VERSION : 0.1
   VAR
      "1#炉体循环水泵电动阀" : "阀门_MODEL";
      "2#炉体循环水泵电动阀" : "阀门_MODEL";
      "3#炉体循环水泵电动阀" : "阀门_MODEL";
      "1#电极循环水泵电动阀" : "阀门_MODEL";
      "2#电极循环水泵电动阀" : "阀门_MODEL";
      "3#电极循环水泵电动阀" : "阀门_MODEL";
      "4#电极循环水泵电动阀" : "阀门_MODEL";
      "1#净环热水泵电动阀" : "阀门_MODEL";
      "2#净环热水泵电动阀" : "阀门_MODEL";
      "3#净环热水泵电动阀" : "阀门_MODEL";
      "4#净环热水泵电动阀" : "阀门_MODEL";
      "5#净环热水泵电动阀" : "阀门_MODEL";
      "1#浊环热水泵电动阀" : "阀门_MODEL";
      "2#浊环热水泵电动阀" : "阀门_MODEL";
      "3#浊环热水泵电动阀" : "阀门_MODEL";
      "4#浊环热水泵电动阀" : "阀门_MODEL";
      "5#浊环热水泵电动阀" : "阀门_MODEL";
      "6#浊环热水泵电动阀" : "阀门_MODEL";
      "7#浊环热水泵电动阀" : "阀门_MODEL";
      "8#浊环热水泵电动阀" : "阀门_MODEL";
      "1#冲渣泵电动阀" : "阀门_MODEL";
      "2#冲渣泵电动阀" : "阀门_MODEL";
      "3#冲渣泵电动阀" : "阀门_MODEL";
      "4#冲渣泵电动阀" : "阀门_MODEL";
      "5#冲渣泵电动阀" : "阀门_MODEL";
      "6#冲渣泵电动阀" : "阀门_MODEL";
      "7#冲渣泵电动阀" : "阀门_MODEL";
      "8#冲渣泵电动阀" : "阀门_MODEL";
      "1#柴油泵电动阀" : "阀门_MODEL";
      "2#柴油泵电动阀" : "阀门_MODEL";
      窑冷却泵电动阀 : "阀门_MODEL";
      Static4_1 : "阀门_MODEL";
      Static5_1 : "阀门_MODEL";
      Static6_1 : "阀门_MODEL";
      Static7_1 : "阀门_MODEL";
      Static8_1 : "阀门_MODEL";
      Static9_1 : "阀门_MODEL";
      Static10_1 : "阀门_MODEL";
      Static11_1 : "阀门_MODEL";
      Static12_1 : "阀门_MODEL";
      Static13_1 : "阀门_MODEL";
      Static14_1 : "阀门_MODEL";
      Static15_1 : "阀门_MODEL";
      Static16_1 : "阀门_MODEL";
      Static17_1 : "阀门_MODEL";
      Static18_1 : "阀门_MODEL";
      Static19_1 : "阀门_MODEL";
      Static20_1 : "阀门_MODEL";
      Static21_1 : "阀门_MODEL";
      Static22_1 : "阀门_MODEL";
      Static23_1 : "阀门_MODEL";
      Static24_1 : "阀门_MODEL";
      Static25_1 : "阀门_MODEL";
      Static26_1 : "阀门_MODEL";
      Static27_1 : "阀门_MODEL";
      Static28_1 : "阀门_MODEL";
      Static29_1 : "阀门_MODEL";
      Static30_1 : "阀门_MODEL";
      Static31_1 : "阀门_MODEL";
      Static32_1 : "阀门_MODEL";
      Static33_1 : "阀门_MODEL";
      Static34_1 : "阀门_MODEL";
      Static35_1 : "阀门_MODEL";
      Static36_1 : "阀门_MODEL";
      Static37_1 : "阀门_MODEL";
      Static38_1 : "阀门_MODEL";
      Static39_1 : "阀门_MODEL";
      Static40_1 : "阀门_MODEL";
      Static41_1 : "阀门_MODEL";
      Static42_1 : "阀门_MODEL";
      Static43_1 : "阀门_MODEL";
      Static44_1 : "阀门_MODEL";
      Static45_1 : "阀门_MODEL";
      Static46_1 : "阀门_MODEL";
      Static47_1 : "阀门_MODEL";
      Static48_1 : "阀门_MODEL";
      Static49_1 : "阀门_MODEL";
      Static50_1 : "阀门_MODEL";
      Static51_1 : "阀门_MODEL";
      Static52_1 : "阀门_MODEL";
      Static53_1 : "阀门_MODEL";
      Static54_1 : "阀门_MODEL";
      Static55_1 : "阀门_MODEL";
      Static56_1 : "阀门_MODEL";
      Static57_1 : "阀门_MODEL";
      Static58_1 : "阀门_MODEL";
      Static59_1 : "阀门_MODEL";
      Static60_1 : "阀门_MODEL";
      Static61_1 : "阀门_MODEL";
      Static62 : "阀门_MODEL";
      Static63 : "阀门_MODEL";
      Static64 : "阀门_MODEL";
      Static65 : "阀门_MODEL";
      Static66 : "阀门_MODEL";
      Static67 : "阀门_MODEL";
      Static68 : "阀门_MODEL";
      Static69 : "阀门_MODEL";
      Static70 : "阀门_MODEL";
      Static71 : "阀门_MODEL";
      Static72 : "阀门_MODEL";
      Static73 : "阀门_MODEL";
      Static74 : "阀门_MODEL";
      阀门_MODEL_Instance : "阀门_MODEL";
   END_VAR
   VAR CONSTANT
      Static3 : Bool;
      Static4 : Bool;
      Static5 : Bool;
      Static6 : Bool;
      Static7 : Bool;
      Static8 : Bool;
      Static9 : Bool;
      Static10 : Bool;
      Static11 : Bool;
      Static12 : Bool;
      Static13 : Bool;
      Static14 : Bool;
      Static15 : Bool;
      Static16 : Bool;
      Static17 : Bool;
      Static18 : Bool;
      Static19 : Bool;
      Static20 : Bool;
      Static21 : Bool;
      Static22 : Bool;
      Static23 : Bool;
      Static24 : Bool;
      Static25 : Bool;
      Static26 : Bool;
      Static27 : Bool;
      Static28 : Bool;
      Static29 : Bool;
      Static30 : Bool;
      Static31 : Bool;
      Static32 : Bool;
      Static33 : Bool;
      Static34 : Bool;
      Static35 : Bool;
      Static36 : Bool;
      Static37 : Bool;
      Static38 : Bool;
      Static39 : Bool;
      Static40 : Bool;
      Static41 : Bool;
      Static42 : Bool;
      Static43 : Bool;
      Static44 : Bool;
      Static45 : Bool;
      Static46 : Bool;
      Static47 : Bool;
      Static48 : Bool;
      Static49 : Bool;
      Static50 : Bool;
      Static51 : Bool;
      Static52 : Bool;
      Static53 : Bool;
      Static54 : Bool;
      Static55 : Bool;
      Static56 : Bool;
      Static57 : Bool;
      Static58 : Bool;
      Static59 : Bool;
      Static60 : Bool;
      Static61 : Bool;
   END_VAR
BEGIN

REGION Network 1
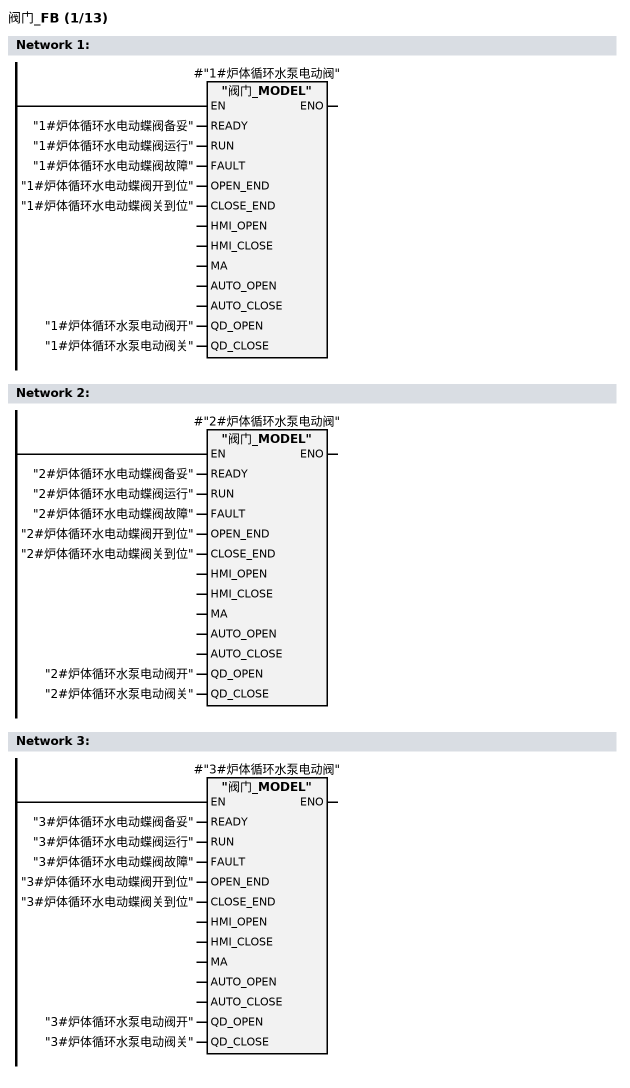
   RUNG wire#powerrail
      #"1#炉体循环水泵电动阀"(READY := "1#炉体循环水电动蝶阀备妥", RUN := "1#炉体循环水电动蝶阀运行", FAULT := "1#炉体循环水电动蝶阀故障", OPEN_END := "1#炉体循环水电动蝶阀开到位", CLOSE_END := "1#炉体循环水电动蝶阀关到位", HMI_OPEN :=, HMI_CLOSE :=, MA :=, AUTO_OPEN :=, AUTO_CLOSE :=, QD_OPEN := "1#炉体循环水泵电动阀开", QD_CLOSE := "1#炉体循环水泵电动阀关")
   END_RUNG
   // the same network as SCL:
   #"1#炉体循环水泵电动阀"(READY := "1#炉体循环水电动蝶阀备妥",   // "阀门_MODEL"
                  RUN := "1#炉体循环水电动蝶阀运行",
                  FAULT := "1#炉体循环水电动蝶阀故障",
                  OPEN_END := "1#炉体循环水电动蝶阀开到位",
                  CLOSE_END := "1#炉体循环水电动蝶阀关到位",
                  QD_OPEN := "1#炉体循环水泵电动阀开",
                  QD_CLOSE := "1#炉体循环水泵电动阀关");
END_REGION

REGION Network 2
   RUNG wire#powerrail
      #"2#炉体循环水泵电动阀"(READY := "2#炉体循环水电动蝶阀备妥", RUN := "2#炉体循环水电动蝶阀运行", FAULT := "2#炉体循环水电动蝶阀故障", OPEN_END := "2#炉体循环水电动蝶阀开到位", CLOSE_END := "2#炉体循环水电动蝶阀关到位", HMI_OPEN :=, HMI_CLOSE :=, MA :=, AUTO_OPEN :=, AUTO_CLOSE :=, QD_OPEN := "2#炉体循环水泵电动阀开", QD_CLOSE := "2#炉体循环水泵电动阀关")
   END_RUNG
   // the same network as SCL:
   #"2#炉体循环水泵电动阀"(READY := "2#炉体循环水电动蝶阀备妥",   // "阀门_MODEL"
                  RUN := "2#炉体循环水电动蝶阀运行",
                  FAULT := "2#炉体循环水电动蝶阀故障",
                  OPEN_END := "2#炉体循环水电动蝶阀开到位",
                  CLOSE_END := "2#炉体循环水电动蝶阀关到位",
                  QD_OPEN := "2#炉体循环水泵电动阀开",
                  QD_CLOSE := "2#炉体循环水泵电动阀关");
END_REGION

REGION Network 3
   RUNG wire#powerrail
      #"3#炉体循环水泵电动阀"(READY := "3#炉体循环水电动蝶阀备妥", RUN := "3#炉体循环水电动蝶阀运行", FAULT := "3#炉体循环水电动蝶阀故障", OPEN_END := "3#炉体循环水电动蝶阀开到位", CLOSE_END := "3#炉体循环水电动蝶阀关到位", HMI_OPEN :=, HMI_CLOSE :=, MA :=, AUTO_OPEN :=, AUTO_CLOSE :=, QD_OPEN := "3#炉体循环水泵电动阀开", QD_CLOSE := "3#炉体循环水泵电动阀关")
   END_RUNG
   // the same network as SCL:
   #"3#炉体循环水泵电动阀"(READY := "3#炉体循环水电动蝶阀备妥",   // "阀门_MODEL"
                  RUN := "3#炉体循环水电动蝶阀运行",
                  FAULT := "3#炉体循环水电动蝶阀故障",
                  OPEN_END := "3#炉体循环水电动蝶阀开到位",
                  CLOSE_END := "3#炉体循环水电动蝶阀关到位",
                  QD_OPEN := "3#炉体循环水泵电动阀开",
                  QD_CLOSE := "3#炉体循环水泵电动阀关");
END_REGION

REGION Network 4
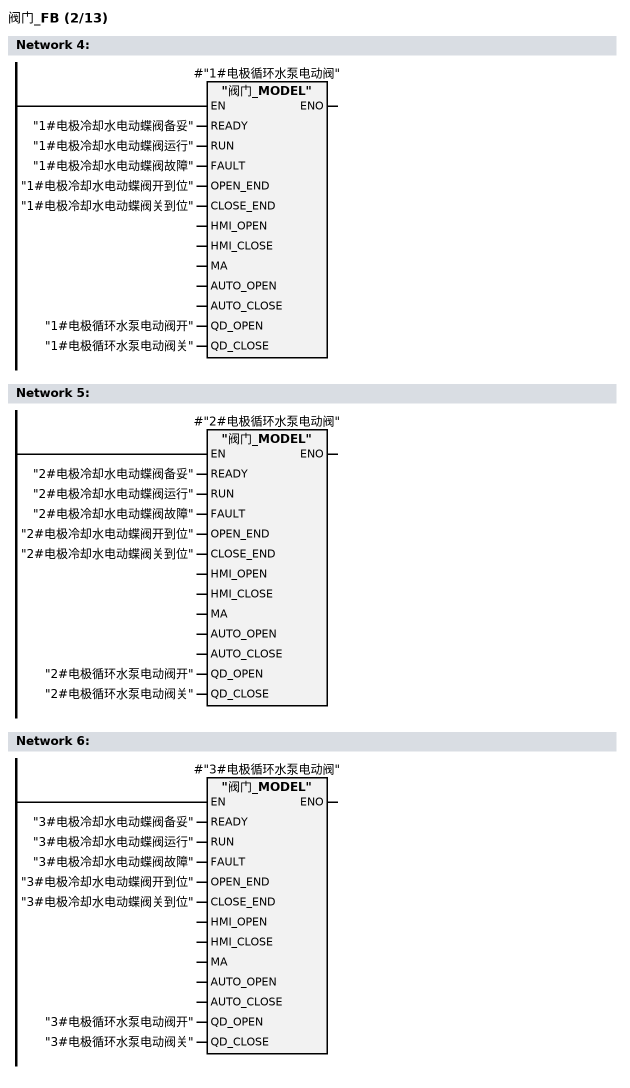
   RUNG wire#powerrail
      #"1#电极循环水泵电动阀"(READY := "1#电极冷却水电动蝶阀备妥", RUN := "1#电极冷却水电动蝶阀运行", FAULT := "1#电极冷却水电动蝶阀故障", OPEN_END := "1#电极冷却水电动蝶阀开到位", CLOSE_END := "1#电极冷却水电动蝶阀关到位", HMI_OPEN :=, HMI_CLOSE :=, MA :=, AUTO_OPEN :=, AUTO_CLOSE :=, QD_OPEN := "1#电极循环水泵电动阀开", QD_CLOSE := "1#电极循环水泵电动阀关")
   END_RUNG
   // the same network as SCL:
   #"1#电极循环水泵电动阀"(READY := "1#电极冷却水电动蝶阀备妥",   // "阀门_MODEL"
                  RUN := "1#电极冷却水电动蝶阀运行",
                  FAULT := "1#电极冷却水电动蝶阀故障",
                  OPEN_END := "1#电极冷却水电动蝶阀开到位",
                  CLOSE_END := "1#电极冷却水电动蝶阀关到位",
                  QD_OPEN := "1#电极循环水泵电动阀开",
                  QD_CLOSE := "1#电极循环水泵电动阀关");
END_REGION

REGION Network 5
   RUNG wire#powerrail
      #"2#电极循环水泵电动阀"(READY := "2#电极冷却水电动蝶阀备妥", RUN := "2#电极冷却水电动蝶阀运行", FAULT := "2#电极冷却水电动蝶阀故障", OPEN_END := "2#电极冷却水电动蝶阀开到位", CLOSE_END := "2#电极冷却水电动蝶阀关到位", HMI_OPEN :=, HMI_CLOSE :=, MA :=, AUTO_OPEN :=, AUTO_CLOSE :=, QD_OPEN := "2#电极循环水泵电动阀开", QD_CLOSE := "2#电极循环水泵电动阀关")
   END_RUNG
   // the same network as SCL:
   #"2#电极循环水泵电动阀"(READY := "2#电极冷却水电动蝶阀备妥",   // "阀门_MODEL"
                  RUN := "2#电极冷却水电动蝶阀运行",
                  FAULT := "2#电极冷却水电动蝶阀故障",
                  OPEN_END := "2#电极冷却水电动蝶阀开到位",
                  CLOSE_END := "2#电极冷却水电动蝶阀关到位",
                  QD_OPEN := "2#电极循环水泵电动阀开",
                  QD_CLOSE := "2#电极循环水泵电动阀关");
END_REGION

REGION Network 6
   RUNG wire#powerrail
      #"3#电极循环水泵电动阀"(READY := "3#电极冷却水电动蝶阀备妥", RUN := "3#电极冷却水电动蝶阀运行", FAULT := "3#电极冷却水电动蝶阀故障", OPEN_END := "3#电极冷却水电动蝶阀开到位", CLOSE_END := "3#电极冷却水电动蝶阀关到位", HMI_OPEN :=, HMI_CLOSE :=, MA :=, AUTO_OPEN :=, AUTO_CLOSE :=, QD_OPEN := "3#电极循环水泵电动阀开", QD_CLOSE := "3#电极循环水泵电动阀关")
   END_RUNG
   // the same network as SCL:
   #"3#电极循环水泵电动阀"(READY := "3#电极冷却水电动蝶阀备妥",   // "阀门_MODEL"
                  RUN := "3#电极冷却水电动蝶阀运行",
                  FAULT := "3#电极冷却水电动蝶阀故障",
                  OPEN_END := "3#电极冷却水电动蝶阀开到位",
                  CLOSE_END := "3#电极冷却水电动蝶阀关到位",
                  QD_OPEN := "3#电极循环水泵电动阀开",
                  QD_CLOSE := "3#电极循环水泵电动阀关");
END_REGION

REGION Network 7
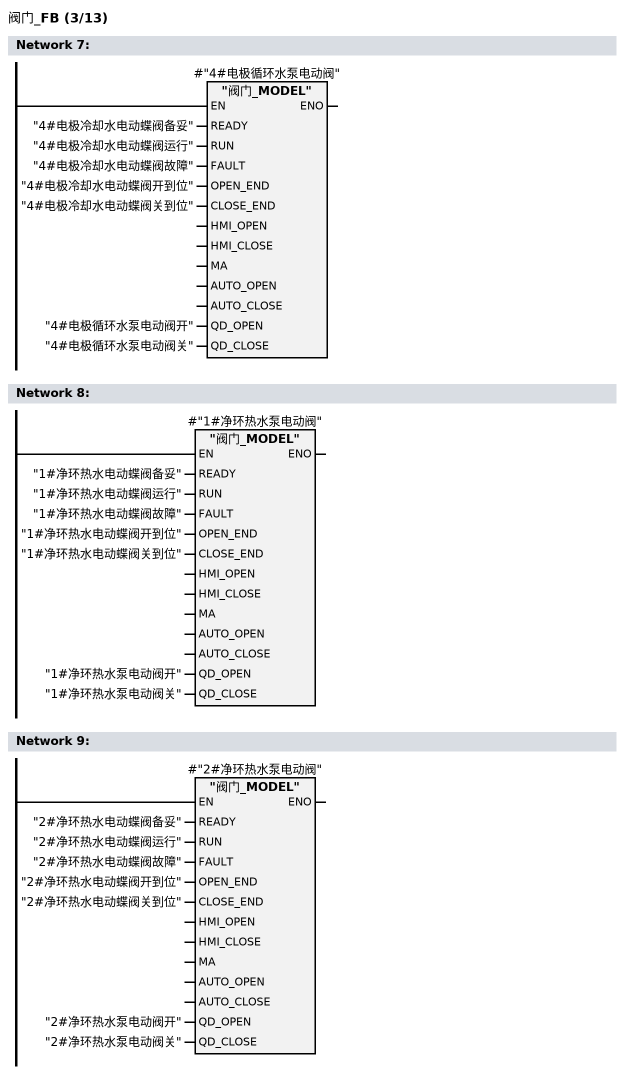
   RUNG wire#powerrail
      #"4#电极循环水泵电动阀"(READY := "4#电极冷却水电动蝶阀备妥", RUN := "4#电极冷却水电动蝶阀运行", FAULT := "4#电极冷却水电动蝶阀故障", OPEN_END := "4#电极冷却水电动蝶阀开到位", CLOSE_END := "4#电极冷却水电动蝶阀关到位", HMI_OPEN :=, HMI_CLOSE :=, MA :=, AUTO_OPEN :=, AUTO_CLOSE :=, QD_OPEN := "4#电极循环水泵电动阀开", QD_CLOSE := "4#电极循环水泵电动阀关")
   END_RUNG
   // the same network as SCL:
   #"4#电极循环水泵电动阀"(READY := "4#电极冷却水电动蝶阀备妥",   // "阀门_MODEL"
                  RUN := "4#电极冷却水电动蝶阀运行",
                  FAULT := "4#电极冷却水电动蝶阀故障",
                  OPEN_END := "4#电极冷却水电动蝶阀开到位",
                  CLOSE_END := "4#电极冷却水电动蝶阀关到位",
                  QD_OPEN := "4#电极循环水泵电动阀开",
                  QD_CLOSE := "4#电极循环水泵电动阀关");
END_REGION

REGION Network 8
   RUNG wire#powerrail
      #"1#净环热水泵电动阀"(READY := "1#净环热水电动蝶阀备妥", RUN := "1#净环热水电动蝶阀运行", FAULT := "1#净环热水电动蝶阀故障", OPEN_END := "1#净环热水电动蝶阀开到位", CLOSE_END := "1#净环热水电动蝶阀关到位", HMI_OPEN :=, HMI_CLOSE :=, MA :=, AUTO_OPEN :=, AUTO_CLOSE :=, QD_OPEN := "1#净环热水泵电动阀开", QD_CLOSE := "1#净环热水泵电动阀关")
   END_RUNG
   // the same network as SCL:
   #"1#净环热水泵电动阀"(READY := "1#净环热水电动蝶阀备妥",   // "阀门_MODEL"
                 RUN := "1#净环热水电动蝶阀运行",
                 FAULT := "1#净环热水电动蝶阀故障",
                 OPEN_END := "1#净环热水电动蝶阀开到位",
                 CLOSE_END := "1#净环热水电动蝶阀关到位",
                 QD_OPEN := "1#净环热水泵电动阀开",
                 QD_CLOSE := "1#净环热水泵电动阀关");
END_REGION

REGION Network 9
   RUNG wire#powerrail
      #"2#净环热水泵电动阀"(READY := "2#净环热水电动蝶阀备妥", RUN := "2#净环热水电动蝶阀运行", FAULT := "2#净环热水电动蝶阀故障", OPEN_END := "2#净环热水电动蝶阀开到位", CLOSE_END := "2#净环热水电动蝶阀关到位", HMI_OPEN :=, HMI_CLOSE :=, MA :=, AUTO_OPEN :=, AUTO_CLOSE :=, QD_OPEN := "2#净环热水泵电动阀开", QD_CLOSE := "2#净环热水泵电动阀关")
   END_RUNG
   // the same network as SCL:
   #"2#净环热水泵电动阀"(READY := "2#净环热水电动蝶阀备妥",   // "阀门_MODEL"
                 RUN := "2#净环热水电动蝶阀运行",
                 FAULT := "2#净环热水电动蝶阀故障",
                 OPEN_END := "2#净环热水电动蝶阀开到位",
                 CLOSE_END := "2#净环热水电动蝶阀关到位",
                 QD_OPEN := "2#净环热水泵电动阀开",
                 QD_CLOSE := "2#净环热水泵电动阀关");
END_REGION

REGION Network 10
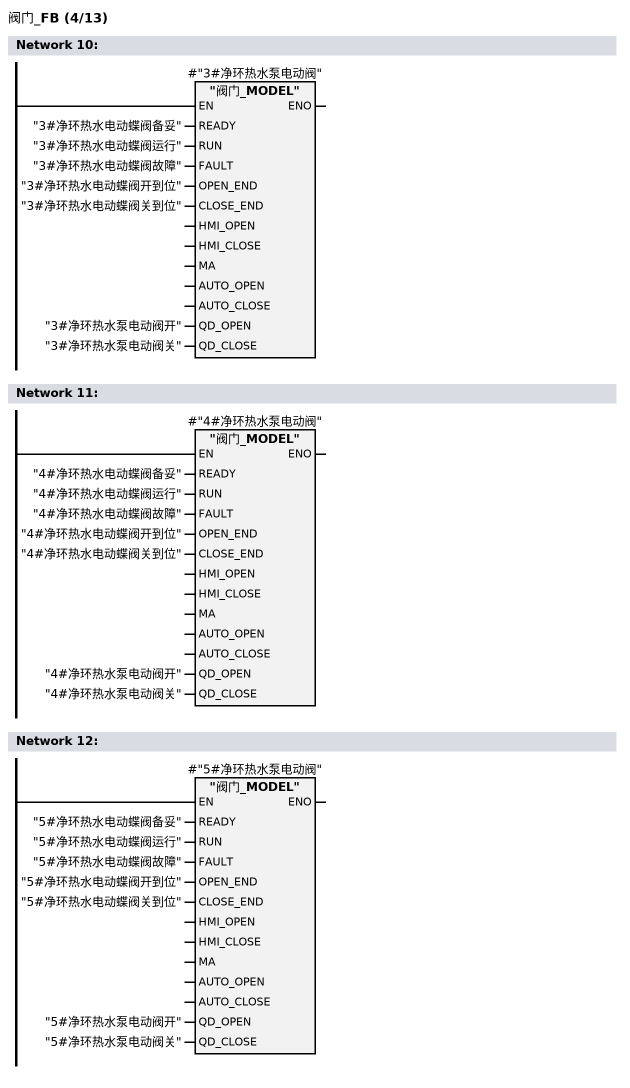
   RUNG wire#powerrail
      #"3#净环热水泵电动阀"(READY := "3#净环热水电动蝶阀备妥", RUN := "3#净环热水电动蝶阀运行", FAULT := "3#净环热水电动蝶阀故障", OPEN_END := "3#净环热水电动蝶阀开到位", CLOSE_END := "3#净环热水电动蝶阀关到位", HMI_OPEN :=, HMI_CLOSE :=, MA :=, AUTO_OPEN :=, AUTO_CLOSE :=, QD_OPEN := "3#净环热水泵电动阀开", QD_CLOSE := "3#净环热水泵电动阀关")
   END_RUNG
   // the same network as SCL:
   #"3#净环热水泵电动阀"(READY := "3#净环热水电动蝶阀备妥",   // "阀门_MODEL"
                 RUN := "3#净环热水电动蝶阀运行",
                 FAULT := "3#净环热水电动蝶阀故障",
                 OPEN_END := "3#净环热水电动蝶阀开到位",
                 CLOSE_END := "3#净环热水电动蝶阀关到位",
                 QD_OPEN := "3#净环热水泵电动阀开",
                 QD_CLOSE := "3#净环热水泵电动阀关");
END_REGION

REGION Network 11
   RUNG wire#powerrail
      #"4#净环热水泵电动阀"(READY := "4#净环热水电动蝶阀备妥", RUN := "4#净环热水电动蝶阀运行", FAULT := "4#净环热水电动蝶阀故障", OPEN_END := "4#净环热水电动蝶阀开到位", CLOSE_END := "4#净环热水电动蝶阀关到位", HMI_OPEN :=, HMI_CLOSE :=, MA :=, AUTO_OPEN :=, AUTO_CLOSE :=, QD_OPEN := "4#净环热水泵电动阀开", QD_CLOSE := "4#净环热水泵电动阀关")
   END_RUNG
   // the same network as SCL:
   #"4#净环热水泵电动阀"(READY := "4#净环热水电动蝶阀备妥",   // "阀门_MODEL"
                 RUN := "4#净环热水电动蝶阀运行",
                 FAULT := "4#净环热水电动蝶阀故障",
                 OPEN_END := "4#净环热水电动蝶阀开到位",
                 CLOSE_END := "4#净环热水电动蝶阀关到位",
                 QD_OPEN := "4#净环热水泵电动阀开",
                 QD_CLOSE := "4#净环热水泵电动阀关");
END_REGION

REGION Network 12
   RUNG wire#powerrail
      #"5#净环热水泵电动阀"(READY := "5#净环热水电动蝶阀备妥", RUN := "5#净环热水电动蝶阀运行", FAULT := "5#净环热水电动蝶阀故障", OPEN_END := "5#净环热水电动蝶阀开到位", CLOSE_END := "5#净环热水电动蝶阀关到位", HMI_OPEN :=, HMI_CLOSE :=, MA :=, AUTO_OPEN :=, AUTO_CLOSE :=, QD_OPEN := "5#净环热水泵电动阀开", QD_CLOSE := "5#净环热水泵电动阀关")
   END_RUNG
   // the same network as SCL:
   #"5#净环热水泵电动阀"(READY := "5#净环热水电动蝶阀备妥",   // "阀门_MODEL"
                 RUN := "5#净环热水电动蝶阀运行",
                 FAULT := "5#净环热水电动蝶阀故障",
                 OPEN_END := "5#净环热水电动蝶阀开到位",
                 CLOSE_END := "5#净环热水电动蝶阀关到位",
                 QD_OPEN := "5#净环热水泵电动阀开",
                 QD_CLOSE := "5#净环热水泵电动阀关");
END_REGION

REGION Network 13
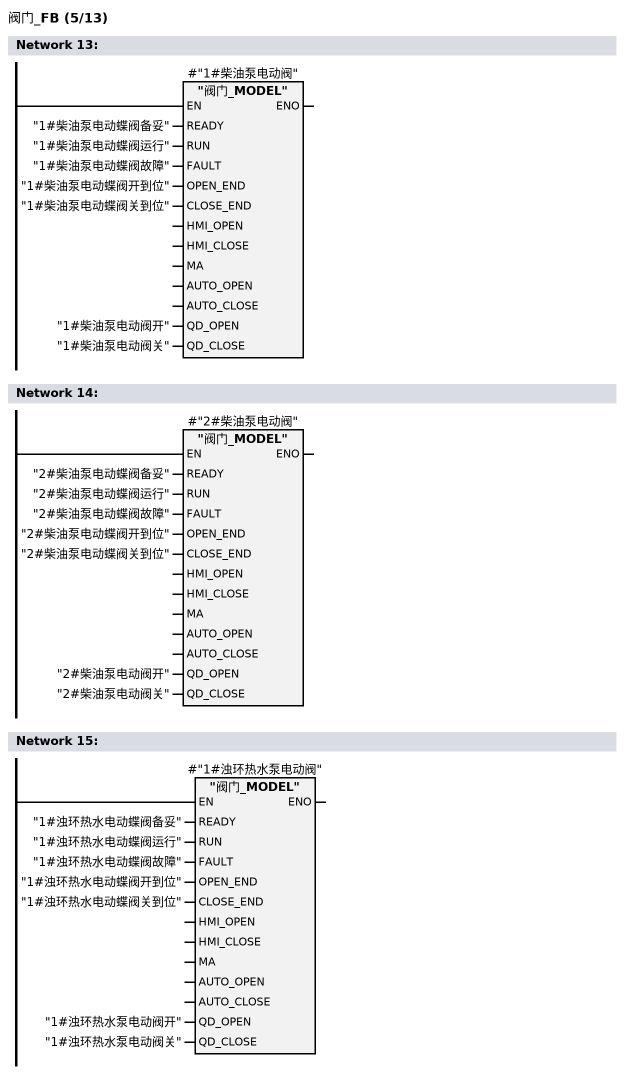
   RUNG wire#powerrail
      #"1#柴油泵电动阀"(READY := "1#柴油泵电动蝶阀备妥", RUN := "1#柴油泵电动蝶阀运行", FAULT := "1#柴油泵电动蝶阀故障", OPEN_END := "1#柴油泵电动蝶阀开到位", CLOSE_END := "1#柴油泵电动蝶阀关到位", HMI_OPEN :=, HMI_CLOSE :=, MA :=, AUTO_OPEN :=, AUTO_CLOSE :=, QD_OPEN := "1#柴油泵电动阀开", QD_CLOSE := "1#柴油泵电动阀关")
   END_RUNG
   // the same network as SCL:
   #"1#柴油泵电动阀"(READY := "1#柴油泵电动蝶阀备妥",   // "阀门_MODEL"
               RUN := "1#柴油泵电动蝶阀运行",
               FAULT := "1#柴油泵电动蝶阀故障",
               OPEN_END := "1#柴油泵电动蝶阀开到位",
               CLOSE_END := "1#柴油泵电动蝶阀关到位",
               QD_OPEN := "1#柴油泵电动阀开",
               QD_CLOSE := "1#柴油泵电动阀关");
END_REGION
